(* Logix 5000 project; controller NWGG 1756-L72 rev 35.12; software revision 35.00; part 16 of 19 *)
(* tags used below, declared in another part *)
   Air_Gates_Opened : BOOL;
   All_Stop : BOOL;
   ALM_K_Valve1_Treat_Failed : ALARM_DIGITAL;
   ALM_KValve0_Clean_Failed : ALARM_DIGITAL;
   ALM_KValve0_Treat_Failed : ALARM_DIGITAL;
   ALM_KValve1_Clean_Failed : ALARM_DIGITAL;
   ALM_OVRAMP_CPLeg : ALARM_DIGITAL;
   ALM_PLUG_CPLeg : ALARM_DIGITAL;
   ALM_SLP10_CPLeg : ALARM_DIGITAL;
   ALM_SLP20_CPLeg : ALARM_DIGITAL;
   ALM_WONT_START_CPLeg : ALARM_DIGITAL;
   Andco_Rate : DINT;
   Auto_Mode : BOOL;
   Auto_Mode_ONS : BOOL;
   Available_For_Clean_Loadout : DINT;
   Available_For_Treat_Loadout : DINT;
   Batch_Status : DINT;
   Belt : udt_Motor[16];
   Belt_Gate_Leg_ON : BOOL;
   Belts_Running : BOOL;
   Bin_Variety_Id : STRING[30];
   Bins_Rqd : BOOL;
   Clean_Batch_Status : DINT;
   Clean_Bin_Gates_Opened : BOOL;
   Clean_K_Relay_Not_Used : BOOL;
   CleanHours : DINT;
   CleanMinuets : DINT;
   CleanSeconds : DINT;
   cntCleanTime : COUNTER;
   Concrete_Leg : udt_Motor;
   Concrete_Leg_Interlock : BOOL;
   ConfigureIndex : DINT;
   ConfirmStop : BOOL;
   Current_Dist_List_IDX : DINT;
   Current_System_Msg_idx : DINT;
   IDX : DINT;
   Loadout_Bin : udt_Loadout_Bin[29];
   Loadout_K_Valve : udt_Loadout_K_Valve[2];
   Loadout_K_Valve_Control : Loadout_K_Valve_Control[2];
   Longest_Clean_Start_IDX : DINT;
   Longest_Clean_Start_Time : DINT;
   Longest_Clean_Stop_IDX : DINT;
   Longest_Clean_Stop_Time : DINT;
   Longest_Treat_Start_IDX : DINT;
   Longest_Treat_Start_Time : DINT;
   Longest_Treat_Stop_IDX : DINT;
   Longest_Treat_Stop_Time : DINT;
   Loop_Idx : DINT;
   Manual_Mode : BOOL;
   Reversing_Belt_Fans : udt_Cyclone;
   System_Status_Msg : STRING;
   System_Status_Msgs : STRING[20];
   TMR_Concrete_Fan : TIMER;
   Transfer_Batch_Status : DINT;
   Treat_Batch_Status : DINT;
   Treater_Loadout : udt_Treater_Loadout;
   _701_K_BYPA : ALIAS FOR I8.1;
   _701_K_TREA : ALIAS FOR I8.0;
   _701K_VALVE : ALIAS FOR O13.10;
   CP_Remote_Leg_In : udt_Motor_Remote_In;
   CP_Remote_Leg_Start : DINT;
   TestOneshot : BOOL;
   testOutput : BOOL;
   TestOutputBit : BOOL;
   testStorageBit : BOOL;
   testTmrOffDelay : TIMER;
   textctr : COUNTER;
(* SeedLoadoutMain, continued *)

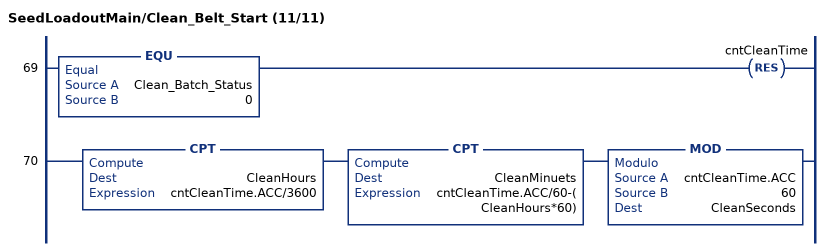
   [picture p317: SeedLoadoutMain/Clean_Belt_Start rungs 69-70]
   69: EQU(Clean_Batch_Status,0)RES(cntCleanTime);
   70: CPT(CleanHours,cntCleanTime.ACC/3600)CPT(CleanMinuets,cntCleanTime.ACC/60-(CleanHours*60))MOD(cntCleanTime.ACC,60,CleanSeconds);
END_ROUTINE

ROUTINE Clean_Bin_Gate_Ready   (* ladder *)
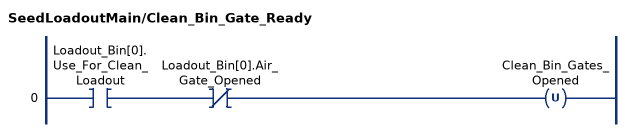
   0: XIC(Loadout_Bin[0].Use_For_Clean_Loadout)XIO(Loadout_Bin[0].Air_Gate_Opened)OTU(Clean_Bin_Gates_Opened);
END_ROUTINE

ROUTINE Clean_Bin_Rqd   (* ladder *)
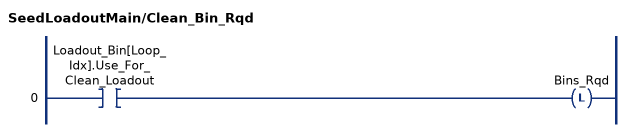
   0: XIC(Loadout_Bin[Loop_Idx].Use_For_Clean_Loadout)OTL(Bins_Rqd);
END_ROUTINE

ROUTINE Close_Air_Gate   (* ladder *)
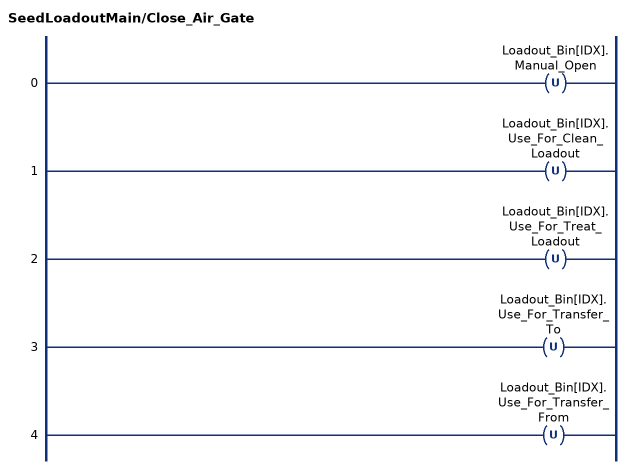
   0: OTU(Loadout_Bin[IDX].Manual_Open);
   1: OTU(Loadout_Bin[IDX].Use_For_Clean_Loadout);
   2: OTU(Loadout_Bin[IDX].Use_For_Treat_Loadout);
   3: OTU(Loadout_Bin[IDX].Use_For_Transfer_To);
   4: OTU(Loadout_Bin[IDX].Use_For_Transfer_From);
END_ROUTINE

ROUTINE Concrete_Leg   (* ladder *)
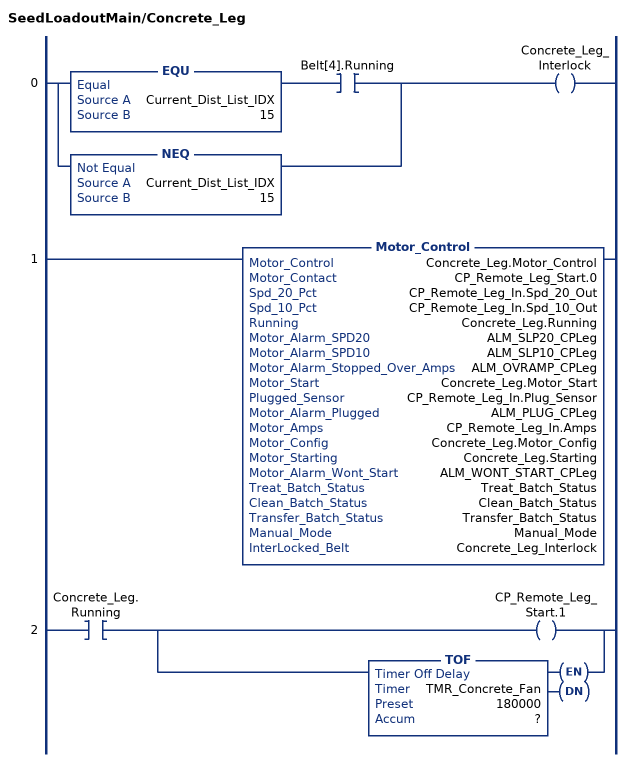
   0: [EQU(Current_Dist_List_IDX,15) XIC(Belt[4].Running) ,NEQ(Current_Dist_List_IDX,15) ]OTE(Concrete_Leg_Interlock);
   1: Motor_Control(Concrete_Leg.Motor_Control,CP_Remote_Leg_Start.0,CP_Remote_Leg_In.Spd_20_Out,CP_Remote_Leg_In.Spd_10_Out,Concrete_Leg.Running,ALM_SLP20_CPLeg,ALM_SLP10_CPLeg,ALM_OVRAMP_CPLeg,Concrete_Leg.Motor_Start,CP_Remote_Leg_In.Plug_Sensor,ALM_PLUG_CPLeg,CP_Remote_Leg_In.Amps,Concrete_Leg.Motor_Config,Concrete_Leg.Starting,ALM_WONT_START_CPLeg,Treat_Batch_Status,Clean_Batch_Status,Transfer_Batch_Status,Manual_Mode,Concrete_Leg_Interlock);
   2: XIC(Concrete_Leg.Running)[OTE(CP_Remote_Leg_Start.1) ,TOF(TMR_Concrete_Fan,?,?) ];
END_ROUTINE

ROUTINE Display   (* ladder *)
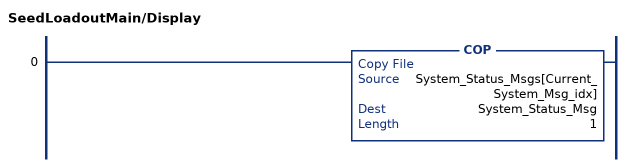
   0: COP(System_Status_Msgs[Current_System_Msg_idx],System_Status_Msg,1);
END_ROUTINE

ROUTINE Get_Longest_Gate_Times   (* ladder *)
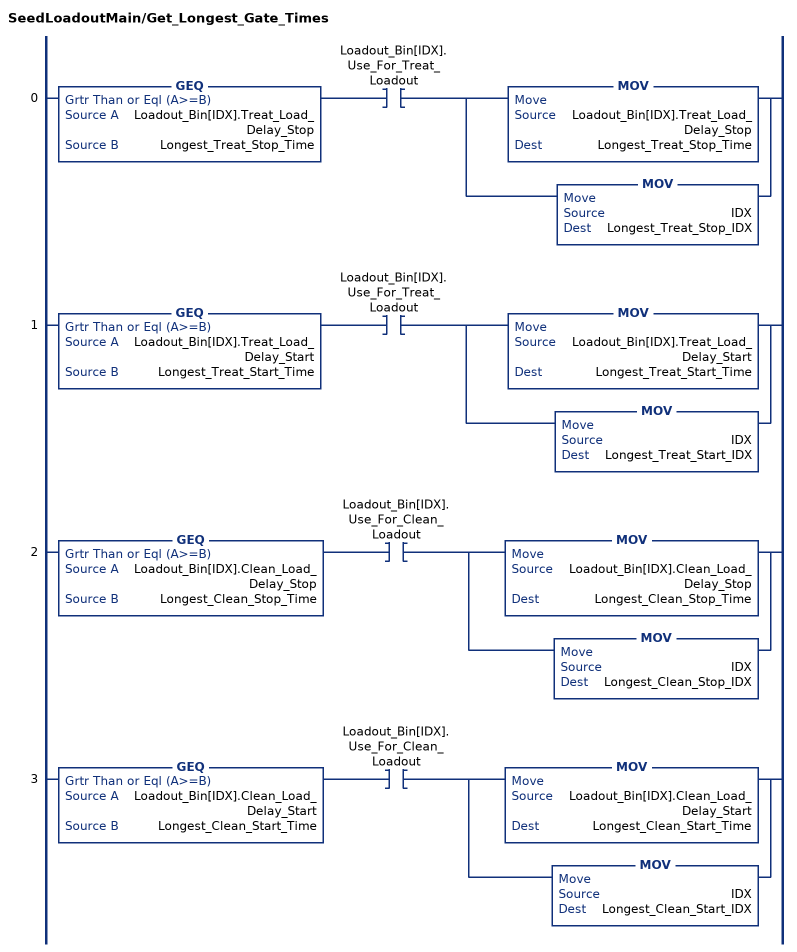
   0: GEQ(Loadout_Bin[IDX].Treat_Load_Delay_Stop,Longest_Treat_Stop_Time)XIC(Loadout_Bin[IDX].Use_For_Treat_Loadout)[MOV(Loadout_Bin[IDX].Treat_Load_Delay_Stop,Longest_Treat_Stop_Time) ,MOV(IDX,Longest_Treat_Stop_IDX) ];
   1: GEQ(Loadout_Bin[IDX].Treat_Load_Delay_Start,Longest_Treat_Start_Time)XIC(Loadout_Bin[IDX].Use_For_Treat_Loadout)[MOV(Loadout_Bin[IDX].Treat_Load_Delay_Start,Longest_Treat_Start_Time) ,MOV(IDX,Longest_Treat_Start_IDX) ];
   2: GEQ(Loadout_Bin[IDX].Clean_Load_Delay_Stop,Longest_Clean_Stop_Time)XIC(Loadout_Bin[IDX].Use_For_Clean_Loadout)[MOV(Loadout_Bin[IDX].Clean_Load_Delay_Stop,Longest_Clean_Stop_Time) ,MOV(IDX,Longest_Clean_Stop_IDX) ];
   3: GEQ(Loadout_Bin[IDX].Clean_Load_Delay_Start,Longest_Clean_Start_Time)XIC(Loadout_Bin[IDX].Use_For_Clean_Loadout)[MOV(Loadout_Bin[IDX].Clean_Load_Delay_Start,Longest_Clean_Start_Time) ,MOV(IDX,Longest_Clean_Start_IDX) ];
END_ROUTINE

ROUTINE Get_System_Status   (* ladder *)
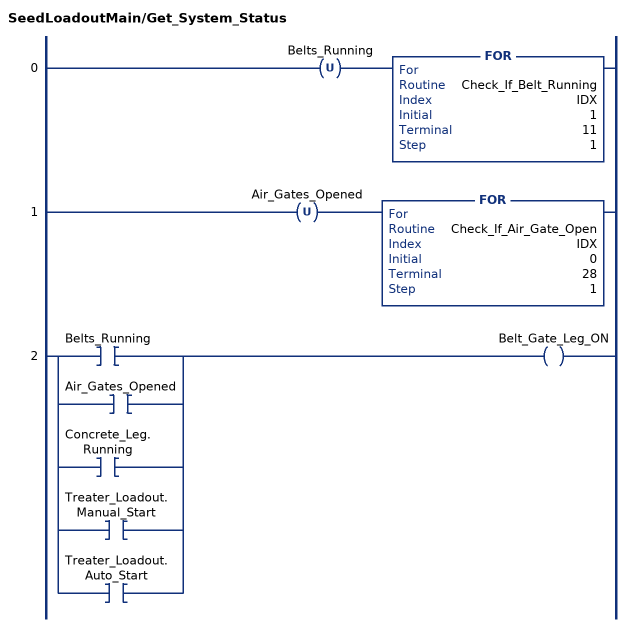
   0: OTU(Belts_Running)FOR(Check_If_Belt_Running,IDX,1,11,1);
   1: OTU(Air_Gates_Opened)FOR(Check_If_Air_Gate_Open,IDX,0,28,1);
   2: [XIC(Belts_Running) ,XIC(Air_Gates_Opened) ,XIC(Concrete_Leg.Running) ,XIC(Treater_Loadout.Manual_Start) ,XIC(Treater_Loadout.Auto_Start) ]OTE(Belt_Gate_Leg_ON);
END_ROUTINE

ROUTINE K_Valves   (* ladder *)
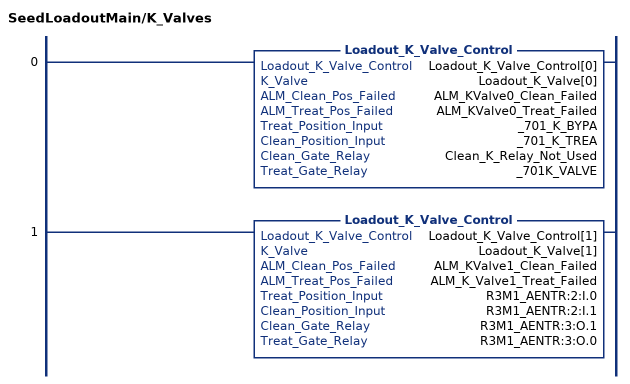
   0: Loadout_K_Valve_Control(Loadout_K_Valve_Control[0],Loadout_K_Valve[0],ALM_KValve0_Clean_Failed,ALM_KValve0_Treat_Failed,_701_K_BYPA,_701_K_TREA,Clean_K_Relay_Not_Used,_701K_VALVE);
   1: Loadout_K_Valve_Control(Loadout_K_Valve_Control[1],Loadout_K_Valve[1],ALM_KValve1_Clean_Failed,ALM_K_Valve1_Treat_Failed,R3M1_AENTR:2:I.0,R3M1_AENTR:2:I.1,R3M1_AENTR:3:O.1,R3M1_AENTR:3:O.0);
END_ROUTINE

ROUTINE Loadout_Time_Delays   (* ladder *)
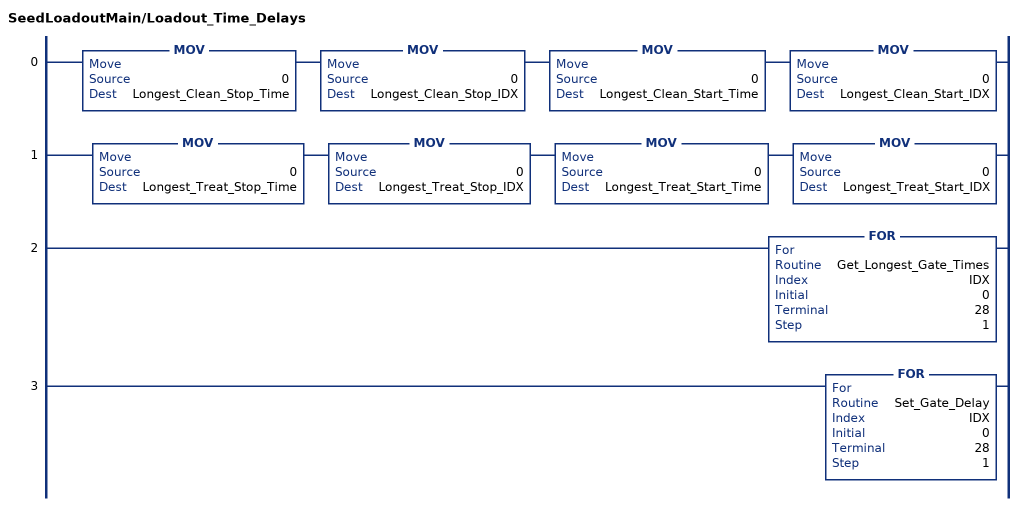
   0: MOV(0,Longest_Clean_Stop_Time)MOV(0,Longest_Clean_Stop_IDX)MOV(0,Longest_Clean_Start_Time)MOV(0,Longest_Clean_Start_IDX);
   1: MOV(0,Longest_Treat_Stop_Time)MOV(0,Longest_Treat_Stop_IDX)MOV(0,Longest_Treat_Start_Time)MOV(0,Longest_Treat_Start_IDX);
   2: FOR(Get_Longest_Gate_Times,IDX,0,28,1);
   3: FOR(Set_Gate_Delay,IDX,0,28,1);
END_ROUTINE

ROUTINE MainRoutine   (* ladder *)
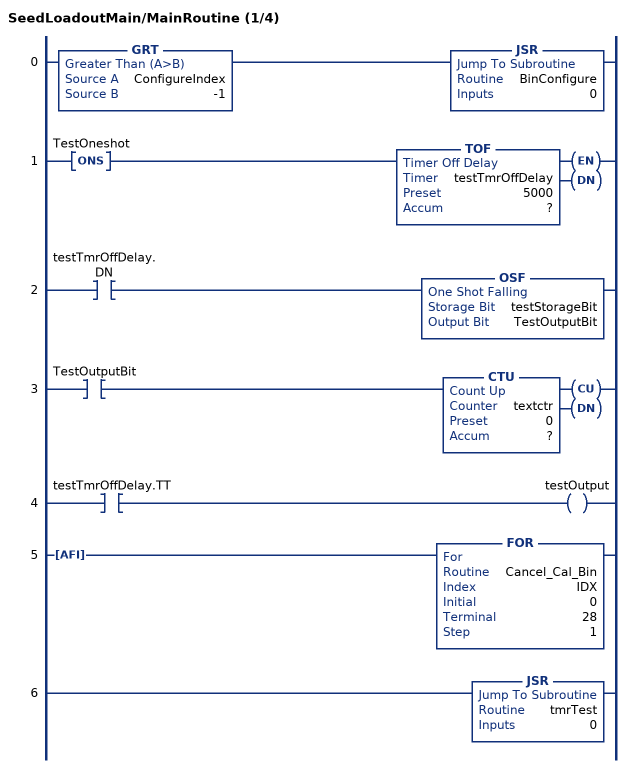
   0: GRT(ConfigureIndex,-1)JSR(BinConfigure,0);
   1: ONS(TestOneshot)TOF(testTmrOffDelay,?,?);
   2: XIC(testTmrOffDelay.DN)OSF(testStorageBit,TestOutputBit);
   3: XIC(TestOutputBit)CTU(textctr,?,?);
   4: XIC(testTmrOffDelay.TT)OTE(testOutput);
   5: AFI()FOR(Cancel_Cal_Bin,IDX,0,28,1);
   6: JSR(tmrTest,0);
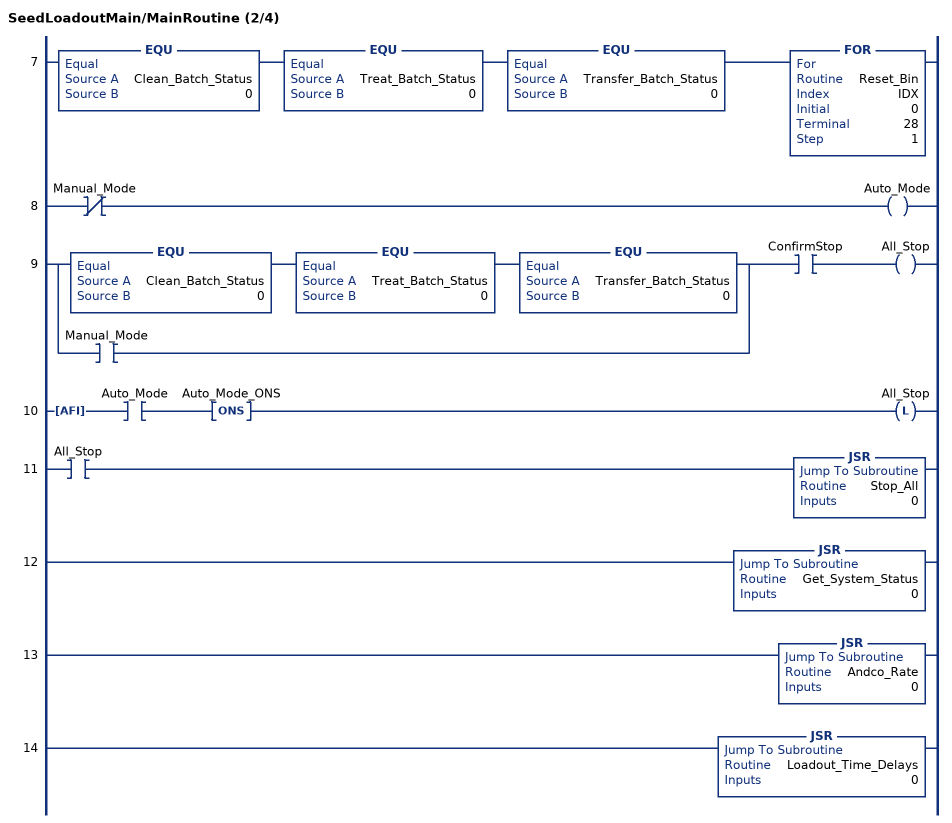
   7: EQU(Clean_Batch_Status,0)EQU(Treat_Batch_Status,0)EQU(Transfer_Batch_Status,0)FOR(Reset_Bin,IDX,0,28,1);
   8: XIO(Manual_Mode)OTE(Auto_Mode);
   9: [EQU(Clean_Batch_Status,0) EQU(Treat_Batch_Status,0) EQU(Transfer_Batch_Status,0) ,XIC(Manual_Mode) ]XIC(ConfirmStop)OTE(All_Stop);
   10: AFI()XIC(Auto_Mode)ONS(Auto_Mode_ONS)OTL(All_Stop);
   11: XIC(All_Stop)JSR(Stop_All,0);
   12: JSR(Get_System_Status,0);
   13: JSR(Andco_Rate,0);
   14: JSR(Loadout_Time_Delays,0);
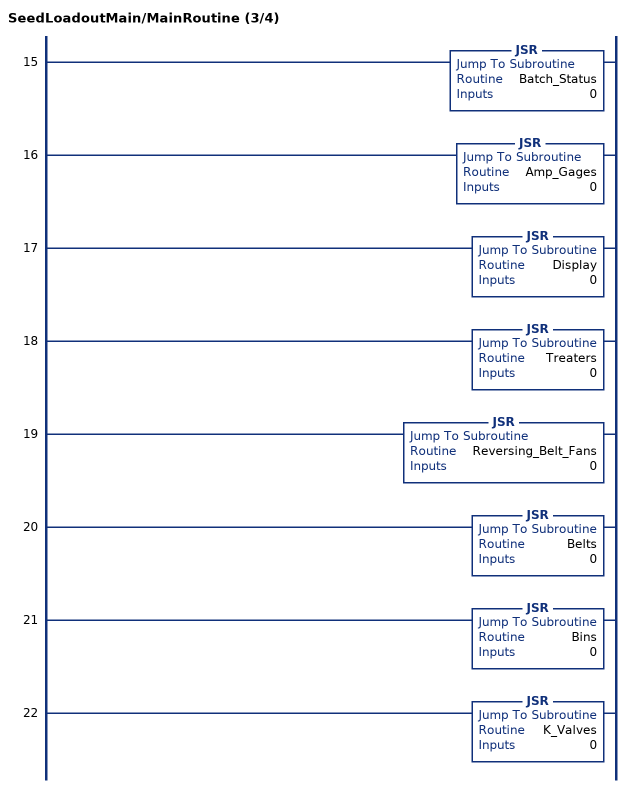
   15: JSR(Batch_Status,0);
   16: JSR(Amp_Gages,0);
   17: JSR(Display,0);
   18: JSR(Treaters,0);
   19: JSR(Reversing_Belt_Fans,0);
   20: JSR(Belts,0);
   21: JSR(Bins,0);
   22: JSR(K_Valves,0);
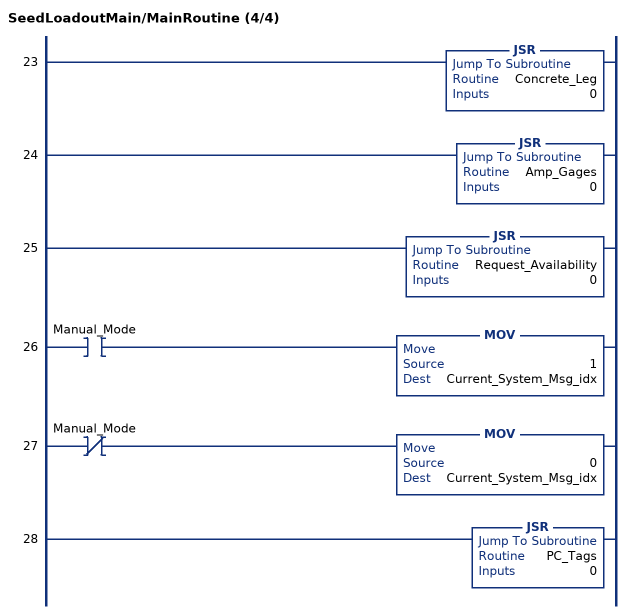
   23: JSR(Concrete_Leg,0);
   24: JSR(Amp_Gages,0);
   25: JSR(Request_Availability,0);
   26: XIC(Manual_Mode)MOV(1,Current_System_Msg_idx);
   27: XIO(Manual_Mode)MOV(0,Current_System_Msg_idx);
   28: JSR(PC_Tags,0);
END_ROUTINE

ROUTINE PC_Tags   (* ladder *)
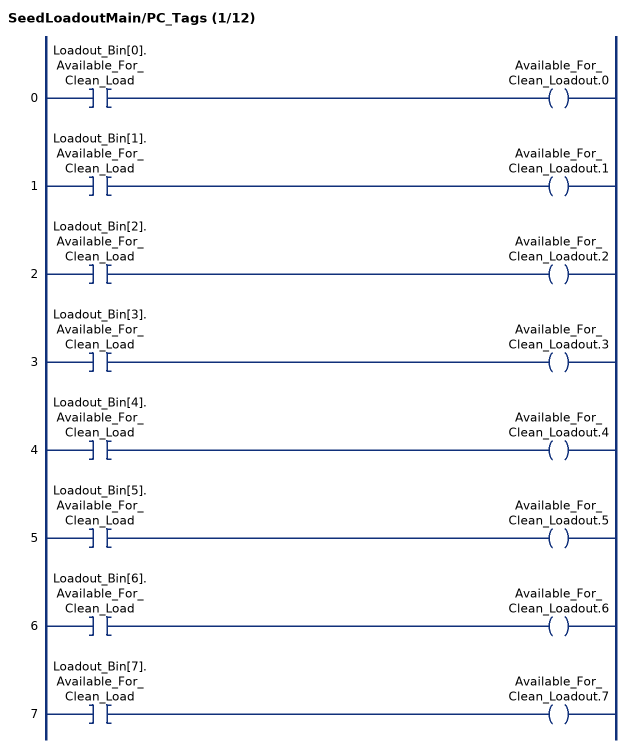
   0: XIC(Loadout_Bin[0].Available_For_Clean_Load)OTE(Available_For_Clean_Loadout.0);
   1: XIC(Loadout_Bin[1].Available_For_Clean_Load)OTE(Available_For_Clean_Loadout.1);
   2: XIC(Loadout_Bin[2].Available_For_Clean_Load)OTE(Available_For_Clean_Loadout.2);
   3: XIC(Loadout_Bin[3].Available_For_Clean_Load)OTE(Available_For_Clean_Loadout.3);
   4: XIC(Loadout_Bin[4].Available_For_Clean_Load)OTE(Available_For_Clean_Loadout.4);
   5: XIC(Loadout_Bin[5].Available_For_Clean_Load)OTE(Available_For_Clean_Loadout.5);
   6: XIC(Loadout_Bin[6].Available_For_Clean_Load)OTE(Available_For_Clean_Loadout.6);
   7: XIC(Loadout_Bin[7].Available_For_Clean_Load)OTE(Available_For_Clean_Loadout.7);
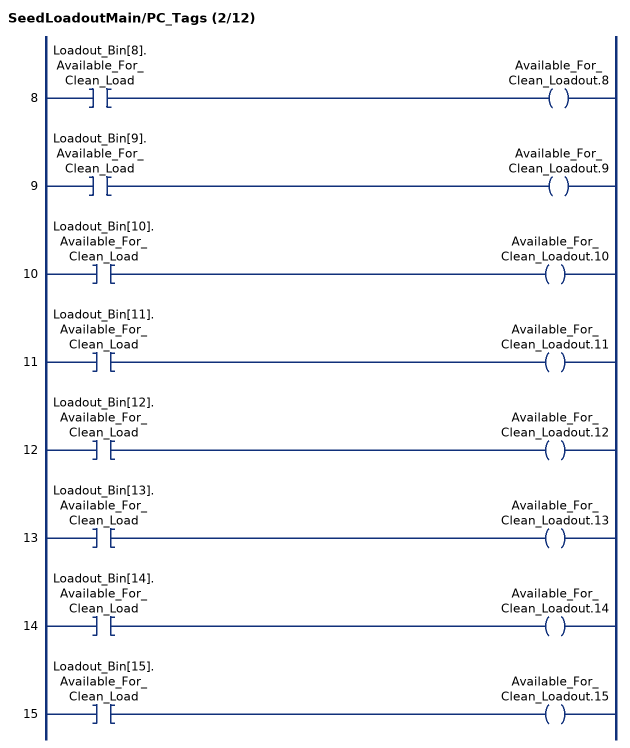
   8: XIC(Loadout_Bin[8].Available_For_Clean_Load)OTE(Available_For_Clean_Loadout.8);
   9: XIC(Loadout_Bin[9].Available_For_Clean_Load)OTE(Available_For_Clean_Loadout.9);
   10: XIC(Loadout_Bin[10].Available_For_Clean_Load)OTE(Available_For_Clean_Loadout.10);
   11: XIC(Loadout_Bin[11].Available_For_Clean_Load)OTE(Available_For_Clean_Loadout.11);
   12: XIC(Loadout_Bin[12].Available_For_Clean_Load)OTE(Available_For_Clean_Loadout.12);
   13: XIC(Loadout_Bin[13].Available_For_Clean_Load)OTE(Available_For_Clean_Loadout.13);
   14: XIC(Loadout_Bin[14].Available_For_Clean_Load)OTE(Available_For_Clean_Loadout.14);
   15: XIC(Loadout_Bin[15].Available_For_Clean_Load)OTE(Available_For_Clean_Loadout.15);
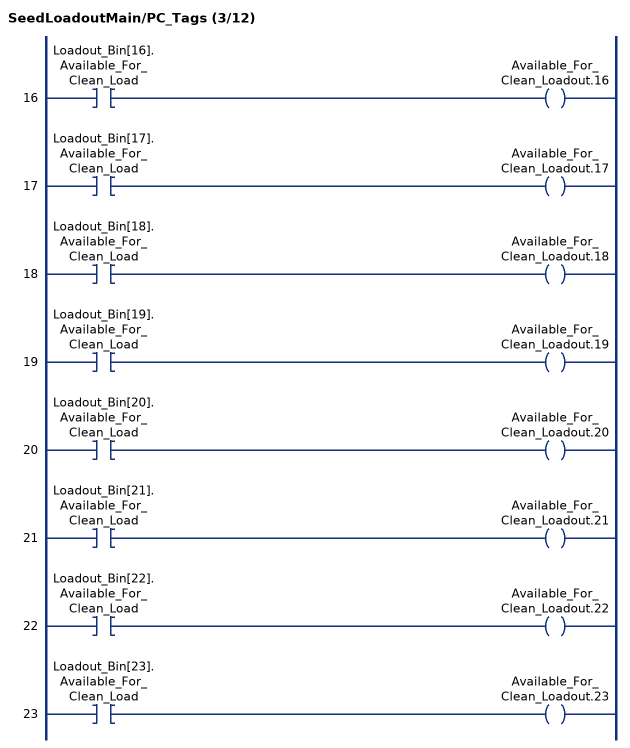
   16: XIC(Loadout_Bin[16].Available_For_Clean_Load)OTE(Available_For_Clean_Loadout.16);
   17: XIC(Loadout_Bin[17].Available_For_Clean_Load)OTE(Available_For_Clean_Loadout.17);
   18: XIC(Loadout_Bin[18].Available_For_Clean_Load)OTE(Available_For_Clean_Loadout.18);
   19: XIC(Loadout_Bin[19].Available_For_Clean_Load)OTE(Available_For_Clean_Loadout.19);
   20: XIC(Loadout_Bin[20].Available_For_Clean_Load)OTE(Available_For_Clean_Loadout.20);
   21: XIC(Loadout_Bin[21].Available_For_Clean_Load)OTE(Available_For_Clean_Loadout.21);
   22: XIC(Loadout_Bin[22].Available_For_Clean_Load)OTE(Available_For_Clean_Loadout.22);
   23: XIC(Loadout_Bin[23].Available_For_Clean_Load)OTE(Available_For_Clean_Loadout.23);
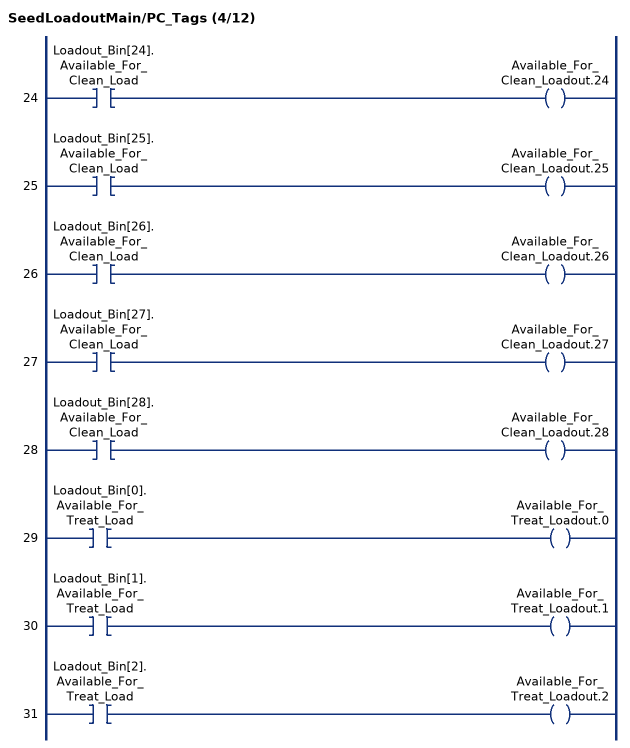
   24: XIC(Loadout_Bin[24].Available_For_Clean_Load)OTE(Available_For_Clean_Loadout.24);
   25: XIC(Loadout_Bin[25].Available_For_Clean_Load)OTE(Available_For_Clean_Loadout.25);
   26: XIC(Loadout_Bin[26].Available_For_Clean_Load)OTE(Available_For_Clean_Loadout.26);
   27: XIC(Loadout_Bin[27].Available_For_Clean_Load)OTE(Available_For_Clean_Loadout.27);
   28: XIC(Loadout_Bin[28].Available_For_Clean_Load)OTE(Available_For_Clean_Loadout.28);
   29: XIC(Loadout_Bin[0].Available_For_Treat_Load)OTE(Available_For_Treat_Loadout.0);
   30: XIC(Loadout_Bin[1].Available_For_Treat_Load)OTE(Available_For_Treat_Loadout.1);
   31: XIC(Loadout_Bin[2].Available_For_Treat_Load)OTE(Available_For_Treat_Loadout.2);
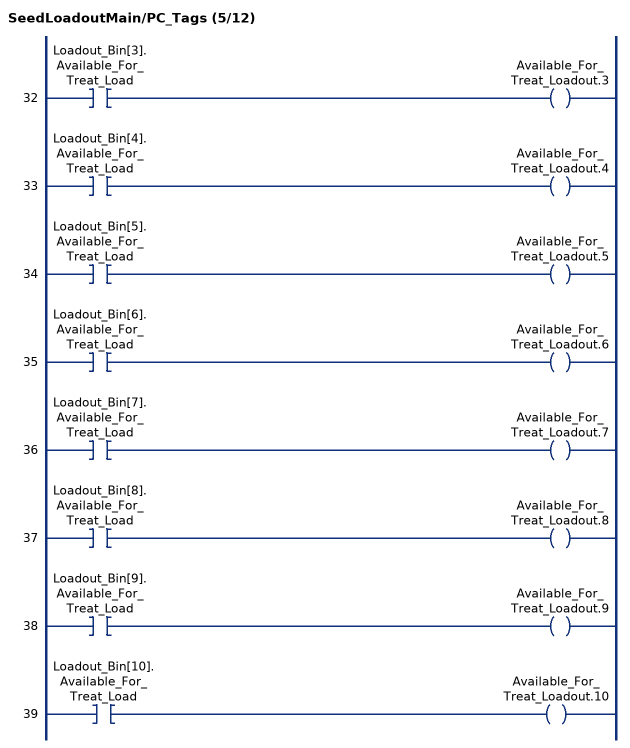
   32: XIC(Loadout_Bin[3].Available_For_Treat_Load)OTE(Available_For_Treat_Loadout.3);
   33: XIC(Loadout_Bin[4].Available_For_Treat_Load)OTE(Available_For_Treat_Loadout.4);
   34: XIC(Loadout_Bin[5].Available_For_Treat_Load)OTE(Available_For_Treat_Loadout.5);
   35: XIC(Loadout_Bin[6].Available_For_Treat_Load)OTE(Available_For_Treat_Loadout.6);
   36: XIC(Loadout_Bin[7].Available_For_Treat_Load)OTE(Available_For_Treat_Loadout.7);
   37: XIC(Loadout_Bin[8].Available_For_Treat_Load)OTE(Available_For_Treat_Loadout.8);
   38: XIC(Loadout_Bin[9].Available_For_Treat_Load)OTE(Available_For_Treat_Loadout.9);
   39: XIC(Loadout_Bin[10].Available_For_Treat_Load)OTE(Available_For_Treat_Loadout.10);
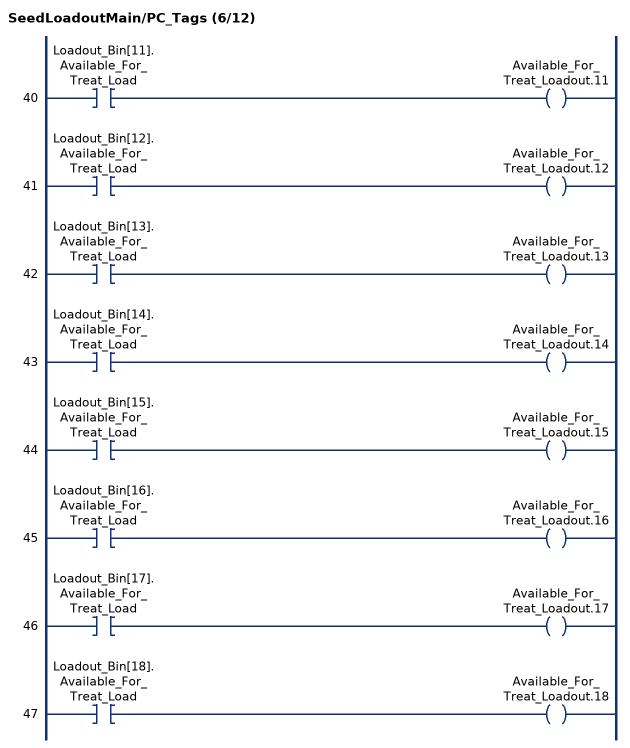
   40: XIC(Loadout_Bin[11].Available_For_Treat_Load)OTE(Available_For_Treat_Loadout.11);
   41: XIC(Loadout_Bin[12].Available_For_Treat_Load)OTE(Available_For_Treat_Loadout.12);
   42: XIC(Loadout_Bin[13].Available_For_Treat_Load)OTE(Available_For_Treat_Loadout.13);
   43: XIC(Loadout_Bin[14].Available_For_Treat_Load)OTE(Available_For_Treat_Loadout.14);
   44: XIC(Loadout_Bin[15].Available_For_Treat_Load)OTE(Available_For_Treat_Loadout.15);
   45: XIC(Loadout_Bin[16].Available_For_Treat_Load)OTE(Available_For_Treat_Loadout.16);
   46: XIC(Loadout_Bin[17].Available_For_Treat_Load)OTE(Available_For_Treat_Loadout.17);
   47: XIC(Loadout_Bin[18].Available_For_Treat_Load)OTE(Available_For_Treat_Loadout.18);
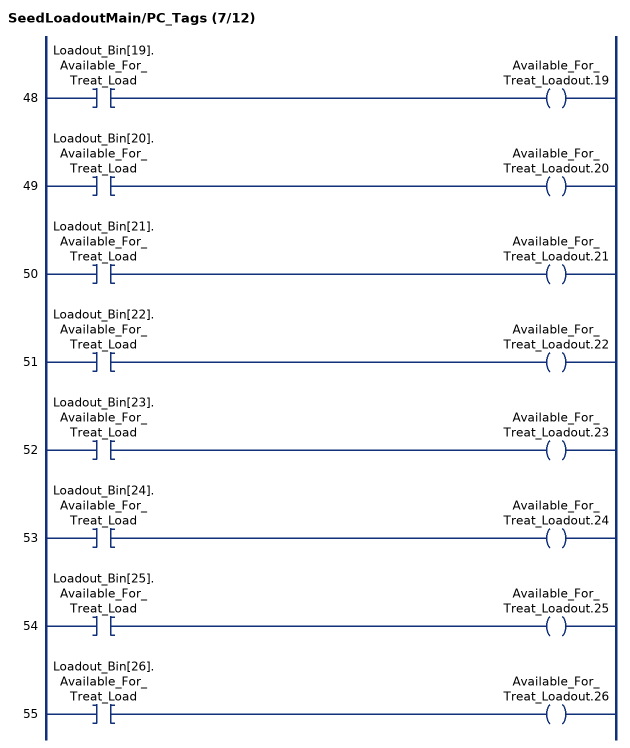
   48: XIC(Loadout_Bin[19].Available_For_Treat_Load)OTE(Available_For_Treat_Loadout.19);
   49: XIC(Loadout_Bin[20].Available_For_Treat_Load)OTE(Available_For_Treat_Loadout.20);
   50: XIC(Loadout_Bin[21].Available_For_Treat_Load)OTE(Available_For_Treat_Loadout.21);
   51: XIC(Loadout_Bin[22].Available_For_Treat_Load)OTE(Available_For_Treat_Loadout.22);
   52: XIC(Loadout_Bin[23].Available_For_Treat_Load)OTE(Available_For_Treat_Loadout.23);
   53: XIC(Loadout_Bin[24].Available_For_Treat_Load)OTE(Available_For_Treat_Loadout.24);
   54: XIC(Loadout_Bin[25].Available_For_Treat_Load)OTE(Available_For_Treat_Loadout.25);
   55: XIC(Loadout_Bin[26].Available_For_Treat_Load)OTE(Available_For_Treat_Loadout.26);
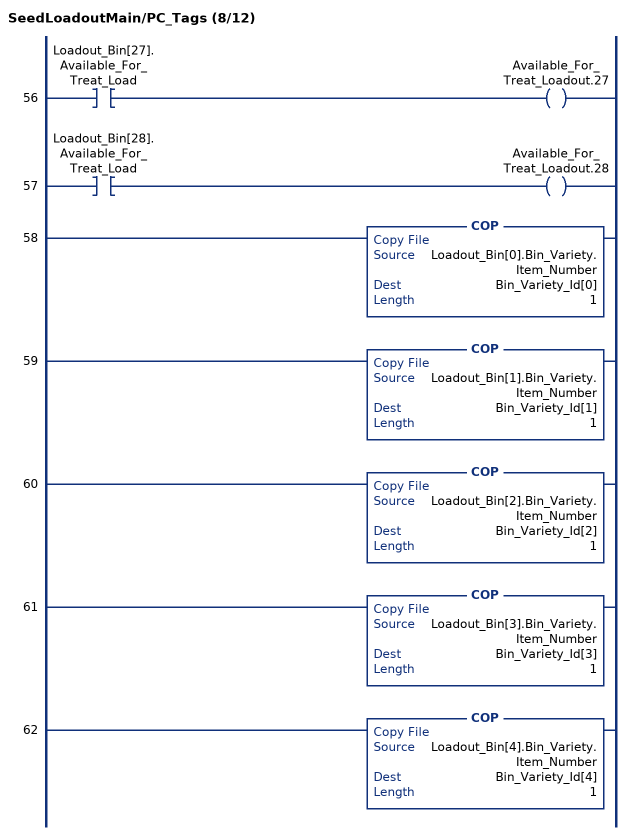
   56: XIC(Loadout_Bin[27].Available_For_Treat_Load)OTE(Available_For_Treat_Loadout.27);
   57: XIC(Loadout_Bin[28].Available_For_Treat_Load)OTE(Available_For_Treat_Loadout.28);
   58: COP(Loadout_Bin[0].Bin_Variety.Item_Number,Bin_Variety_Id[0],1);
   59: COP(Loadout_Bin[1].Bin_Variety.Item_Number,Bin_Variety_Id[1],1);
   60: COP(Loadout_Bin[2].Bin_Variety.Item_Number,Bin_Variety_Id[2],1);
   61: COP(Loadout_Bin[3].Bin_Variety.Item_Number,Bin_Variety_Id[3],1);
   62: COP(Loadout_Bin[4].Bin_Variety.Item_Number,Bin_Variety_Id[4],1);
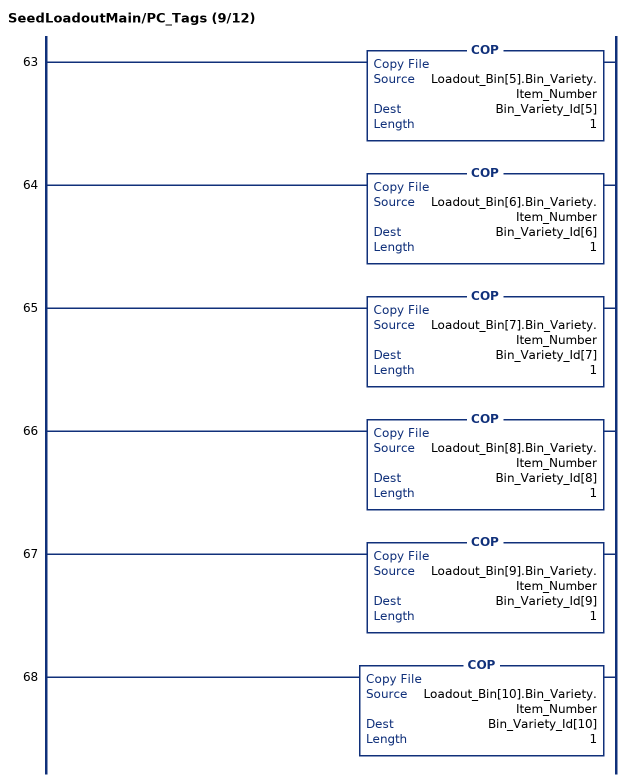
   63: COP(Loadout_Bin[5].Bin_Variety.Item_Number,Bin_Variety_Id[5],1);
   64: COP(Loadout_Bin[6].Bin_Variety.Item_Number,Bin_Variety_Id[6],1);
   65: COP(Loadout_Bin[7].Bin_Variety.Item_Number,Bin_Variety_Id[7],1);
   66: COP(Loadout_Bin[8].Bin_Variety.Item_Number,Bin_Variety_Id[8],1);
   67: COP(Loadout_Bin[9].Bin_Variety.Item_Number,Bin_Variety_Id[9],1);
   68: COP(Loadout_Bin[10].Bin_Variety.Item_Number,Bin_Variety_Id[10],1);
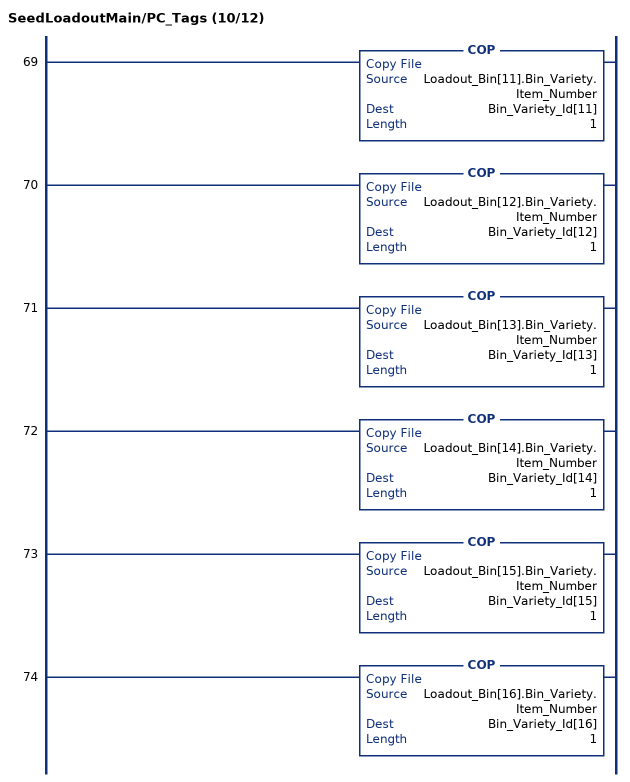
   69: COP(Loadout_Bin[11].Bin_Variety.Item_Number,Bin_Variety_Id[11],1);
   70: COP(Loadout_Bin[12].Bin_Variety.Item_Number,Bin_Variety_Id[12],1);
   71: COP(Loadout_Bin[13].Bin_Variety.Item_Number,Bin_Variety_Id[13],1);
   72: COP(Loadout_Bin[14].Bin_Variety.Item_Number,Bin_Variety_Id[14],1);
   73: COP(Loadout_Bin[15].Bin_Variety.Item_Number,Bin_Variety_Id[15],1);
   74: COP(Loadout_Bin[16].Bin_Variety.Item_Number,Bin_Variety_Id[16],1);
